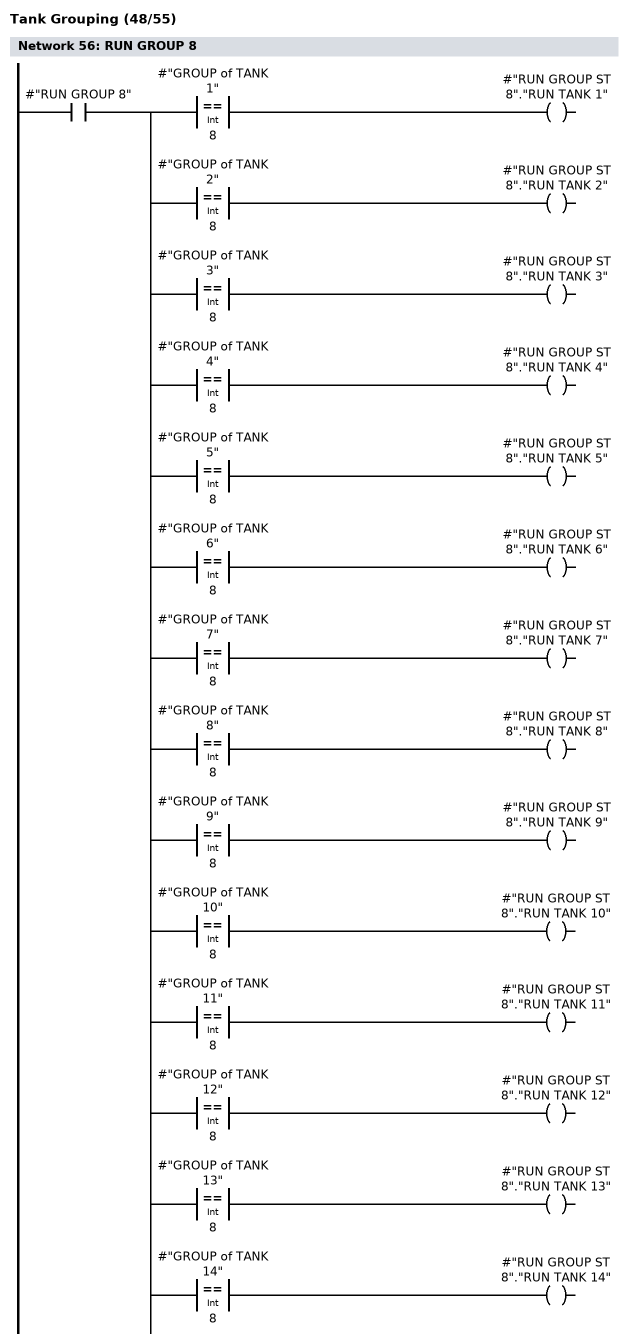
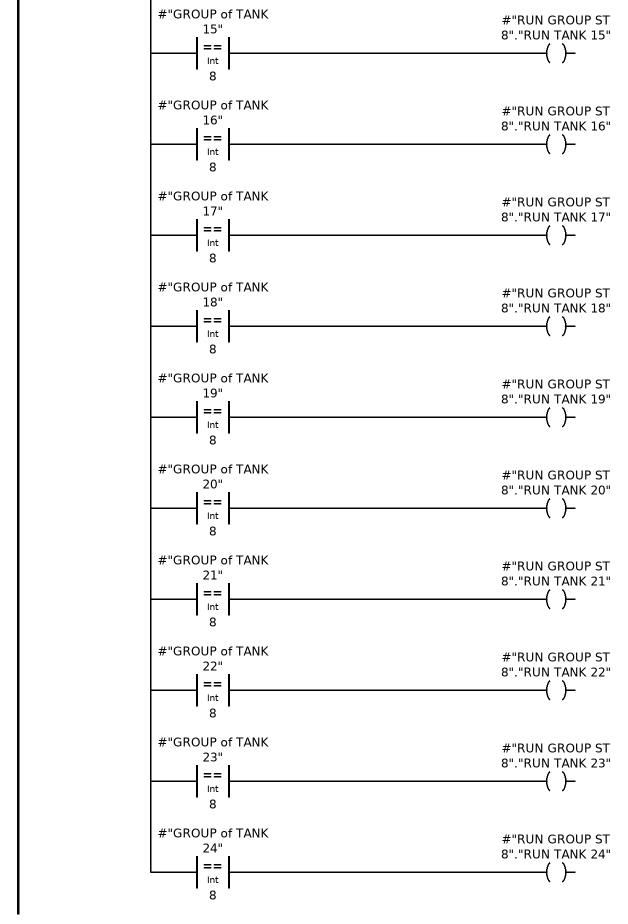
   RUNG wire#powerrail
      Contact( #"RUN GROUP 8" )
      wire#w1
      { S7_Templates := "SrcType := Int" } EQ_Contact(in1 := #"GROUP of TANK 1", in2 := 8)
      Coil( #"RUN GROUP ST 8"."RUN TANK 1" )
   END_RUNG
   RUNG wire#w1
      { S7_Templates := "SrcType := Int" } EQ_Contact(in1 := #"GROUP of TANK 2", in2 := 8)
      Coil( #"RUN GROUP ST 8"."RUN TANK 2" )
   END_RUNG
   RUNG wire#w1
      { S7_Templates := "SrcType := Int" } EQ_Contact(in1 := #"GROUP of TANK 3", in2 := 8)
      Coil( #"RUN GROUP ST 8"."RUN TANK 3" )
   END_RUNG
   RUNG wire#w1
      { S7_Templates := "SrcType := Int" } EQ_Contact(in1 := #"GROUP of TANK 4", in2 := 8)
      Coil( #"RUN GROUP ST 8"."RUN TANK 4" )
   END_RUNG
   RUNG wire#w1
      { S7_Templates := "SrcType := Int" } EQ_Contact(in1 := #"GROUP of TANK 5", in2 := 8)
      Coil( #"RUN GROUP ST 8"."RUN TANK 5" )
   END_RUNG
   RUNG wire#w1
      { S7_Templates := "SrcType := Int" } EQ_Contact(in1 := #"GROUP of TANK 6", in2 := 8)
      Coil( #"RUN GROUP ST 8"."RUN TANK 6" )
   END_RUNG
   RUNG wire#w1
      { S7_Templates := "SrcType := Int" } EQ_Contact(in1 := #"GROUP of TANK 7", in2 := 8)
      Coil( #"RUN GROUP ST 8"."RUN TANK 7" )
   END_RUNG
   RUNG wire#w1
      { S7_Templates := "SrcType := Int" } EQ_Contact(in1 := #"GROUP of TANK 8", in2 := 8)
      Coil( #"RUN GROUP ST 8"."RUN TANK 8" )
   END_RUNG
   RUNG wire#w1
      { S7_Templates := "SrcType := Int" } EQ_Contact(in1 := #"GROUP of TANK 9", in2 := 8)
      Coil( #"RUN GROUP ST 8"."RUN TANK 9" )
   END_RUNG
   RUNG wire#w1
      { S7_Templates := "SrcType := Int" } EQ_Contact(in1 := #"GROUP of TANK 10", in2 := 8)
      Coil( #"RUN GROUP ST 8"."RUN TANK 10" )
   END_RUNG
   RUNG wire#w1
      { S7_Templates := "SrcType := Int" } EQ_Contact(in1 := #"GROUP of TANK 11", in2 := 8)
      Coil( #"RUN GROUP ST 8"."RUN TANK 11" )
   END_RUNG
   RUNG wire#w1
      { S7_Templates := "SrcType := Int" } EQ_Contact(in1 := #"GROUP of TANK 12", in2 := 8)
      Coil( #"RUN GROUP ST 8"."RUN TANK 12" )
   END_RUNG
   RUNG wire#w1
      { S7_Templates := "SrcType := Int" } EQ_Contact(in1 := #"GROUP of TANK 13", in2 := 8)
      Coil( #"RUN GROUP ST 8"."RUN TANK 13" )
   END_RUNG
   RUNG wire#w1
      { S7_Templates := "SrcType := Int" } EQ_Contact(in1 := #"GROUP of TANK 14", in2 := 8)
      Coil( #"RUN GROUP ST 8"."RUN TANK 14" )
   END_RUNG
   RUNG wire#w1
      { S7_Templates := "SrcType := Int" } EQ_Contact(in1 := #"GROUP of TANK 15", in2 := 8)
      Coil( #"RUN GROUP ST 8"."RUN TANK 15" )
   END_RUNG
   RUNG wire#w1
      { S7_Templates := "SrcType := Int" } EQ_Contact(in1 := #"GROUP of TANK 16", in2 := 8)
      Coil( #"RUN GROUP ST 8"."RUN TANK 16" )
   END_RUNG
   RUNG wire#w1
      { S7_Templates := "SrcType := Int" } EQ_Contact(in1 := #"GROUP of TANK 17", in2 := 8)
      Coil( #"RUN GROUP ST 8"."RUN TANK 17" )
   END_RUNG
   RUNG wire#w1
      { S7_Templates := "SrcType := Int" } EQ_Contact(in1 := #"GROUP of TANK 18", in2 := 8)
      Coil( #"RUN GROUP ST 8"."RUN TANK 18" )
   END_RUNG
   RUNG wire#w1
      { S7_Templates := "SrcType := Int" } EQ_Contact(in1 := #"GROUP of TANK 19", in2 := 8)
      Coil( #"RUN GROUP ST 8"."RUN TANK 19" )
   END_RUNG
   RUNG wire#w1
      { S7_Templates := "SrcType := Int" } EQ_Contact(in1 := #"GROUP of TANK 20", in2 := 8)
      Coil( #"RUN GROUP ST 8"."RUN TANK 20" )
   END_RUNG
   RUNG wire#w1
      { S7_Templates := "SrcType := Int" } EQ_Contact(in1 := #"GROUP of TANK 21", in2 := 8)
      Coil( #"RUN GROUP ST 8"."RUN TANK 21" )
   END_RUNG
   RUNG wire#w1
      { S7_Templates := "SrcType := Int" } EQ_Contact(in1 := #"GROUP of TANK 22", in2 := 8)
      Coil( #"RUN GROUP ST 8"."RUN TANK 22" )
   END_RUNG
   RUNG wire#w1
      { S7_Templates := "SrcType := Int" } EQ_Contact(in1 := #"GROUP of TANK 23", in2 := 8)
      Coil( #"RUN GROUP ST 8"."RUN TANK 23" )
   END_RUNG
   RUNG wire#w1
      { S7_Templates := "SrcType := Int" } EQ_Contact(in1 := #"GROUP of TANK 24", in2 := 8)
      Coil( #"RUN GROUP ST 8"."RUN TANK 24" )
   END_RUNG
   // the same network as SCL:
   #"RUN GROUP ST 8"."RUN TANK 1" := #"RUN GROUP 8" AND (#"GROUP of TANK 1" = 8);
   #"RUN GROUP ST 8"."RUN TANK 2" := #"RUN GROUP 8" AND (#"GROUP of TANK 2" = 8);
   #"RUN GROUP ST 8"."RUN TANK 3" := #"RUN GROUP 8" AND (#"GROUP of TANK 3" = 8);
   #"RUN GROUP ST 8"."RUN TANK 4" := #"RUN GROUP 8" AND (#"GROUP of TANK 4" = 8);
   #"RUN GROUP ST 8"."RUN TANK 5" := #"RUN GROUP 8" AND (#"GROUP of TANK 5" = 8);
   #"RUN GROUP ST 8"."RUN TANK 6" := #"RUN GROUP 8" AND (#"GROUP of TANK 6" = 8);
   #"RUN GROUP ST 8"."RUN TANK 7" := #"RUN GROUP 8" AND (#"GROUP of TANK 7" = 8);
   #"RUN GROUP ST 8"."RUN TANK 8" := #"RUN GROUP 8" AND (#"GROUP of TANK 8" = 8);
   #"RUN GROUP ST 8"."RUN TANK 9" := #"RUN GROUP 8" AND (#"GROUP of TANK 9" = 8);
   #"RUN GROUP ST 8"."RUN TANK 10" := #"RUN GROUP 8" AND (#"GROUP of TANK 10" = 8);
   #"RUN GROUP ST 8"."RUN TANK 11" := #"RUN GROUP 8" AND (#"GROUP of TANK 11" = 8);
   #"RUN GROUP ST 8"."RUN TANK 12" := #"RUN GROUP 8" AND (#"GROUP of TANK 12" = 8);
   #"RUN GROUP ST 8"."RUN TANK 13" := #"RUN GROUP 8" AND (#"GROUP of TANK 13" = 8);
   #"RUN GROUP ST 8"."RUN TANK 14" := #"RUN GROUP 8" AND (#"GROUP of TANK 14" = 8);
   #"RUN GROUP ST 8"."RUN TANK 15" := #"RUN GROUP 8" AND (#"GROUP of TANK 15" = 8);
   #"RUN GROUP ST 8"."RUN TANK 16" := #"RUN GROUP 8" AND (#"GROUP of TANK 16" = 8);
   #"RUN GROUP ST 8"."RUN TANK 17" := #"RUN GROUP 8" AND (#"GROUP of TANK 17" = 8);
   #"RUN GROUP ST 8"."RUN TANK 18" := #"RUN GROUP 8" AND (#"GROUP of TANK 18" = 8);
   #"RUN GROUP ST 8"."RUN TANK 19" := #"RUN GROUP 8" AND (#"GROUP of TANK 19" = 8);
   #"RUN GROUP ST 8"."RUN TANK 20" := #"RUN GROUP 8" AND (#"GROUP of TANK 20" = 8);
   #"RUN GROUP ST 8"."RUN TANK 21" := #"RUN GROUP 8" AND (#"GROUP of TANK 21" = 8);
   #"RUN GROUP ST 8"."RUN TANK 22" := #"RUN GROUP 8" AND (#"GROUP of TANK 22" = 8);
   #"RUN GROUP ST 8"."RUN TANK 23" := #"RUN GROUP 8" AND (#"GROUP of TANK 23" = 8);
   #"RUN GROUP ST 8"."RUN TANK 24" := #"RUN GROUP 8" AND (#"GROUP of TANK 24" = 8);
END_REGION

REGION Network 57: RUN GROUP 9
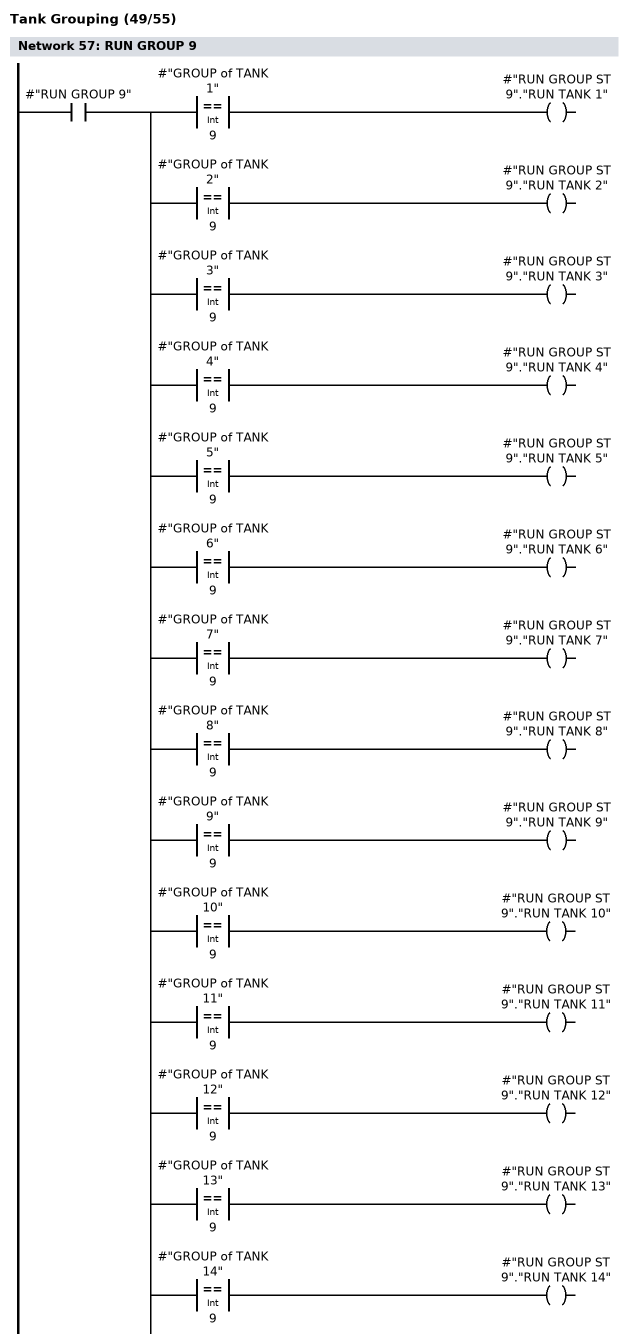
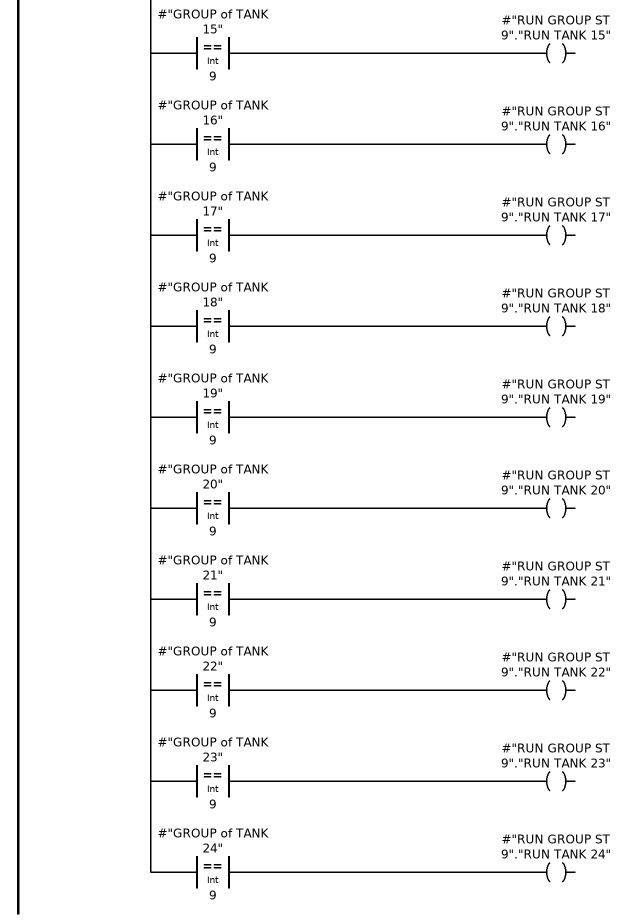
   RUNG wire#powerrail
      Contact( #"RUN GROUP 9" )
      wire#w1
      { S7_Templates := "SrcType := Int" } EQ_Contact(in1 := #"GROUP of TANK 1", in2 := 9)
      Coil( #"RUN GROUP ST 9"."RUN TANK 1" )
   END_RUNG
   RUNG wire#w1
      { S7_Templates := "SrcType := Int" } EQ_Contact(in1 := #"GROUP of TANK 2", in2 := 9)
      Coil( #"RUN GROUP ST 9"."RUN TANK 2" )
   END_RUNG
   RUNG wire#w1
      { S7_Templates := "SrcType := Int" } EQ_Contact(in1 := #"GROUP of TANK 3", in2 := 9)
      Coil( #"RUN GROUP ST 9"."RUN TANK 3" )
   END_RUNG
   RUNG wire#w1
      { S7_Templates := "SrcType := Int" } EQ_Contact(in1 := #"GROUP of TANK 4", in2 := 9)
      Coil( #"RUN GROUP ST 9"."RUN TANK 4" )
   END_RUNG
   RUNG wire#w1
      { S7_Templates := "SrcType := Int" } EQ_Contact(in1 := #"GROUP of TANK 5", in2 := 9)
      Coil( #"RUN GROUP ST 9"."RUN TANK 5" )
   END_RUNG
   RUNG wire#w1
      { S7_Templates := "SrcType := Int" } EQ_Contact(in1 := #"GROUP of TANK 6", in2 := 9)
      Coil( #"RUN GROUP ST 9"."RUN TANK 6" )
   END_RUNG
   RUNG wire#w1
      { S7_Templates := "SrcType := Int" } EQ_Contact(in1 := #"GROUP of TANK 7", in2 := 9)
      Coil( #"RUN GROUP ST 9"."RUN TANK 7" )
   END_RUNG
   RUNG wire#w1
      { S7_Templates := "SrcType := Int" } EQ_Contact(in1 := #"GROUP of TANK 8", in2 := 9)
      Coil( #"RUN GROUP ST 9"."RUN TANK 8" )
   END_RUNG
   RUNG wire#w1
      { S7_Templates := "SrcType := Int" } EQ_Contact(in1 := #"GROUP of TANK 9", in2 := 9)
      Coil( #"RUN GROUP ST 9"."RUN TANK 9" )
   END_RUNG
   RUNG wire#w1
      { S7_Templates := "SrcType := Int" } EQ_Contact(in1 := #"GROUP of TANK 10", in2 := 9)
      Coil( #"RUN GROUP ST 9"."RUN TANK 10" )
   END_RUNG
   RUNG wire#w1
      { S7_Templates := "SrcType := Int" } EQ_Contact(in1 := #"GROUP of TANK 11", in2 := 9)
      Coil( #"RUN GROUP ST 9"."RUN TANK 11" )
   END_RUNG
   RUNG wire#w1
      { S7_Templates := "SrcType := Int" } EQ_Contact(in1 := #"GROUP of TANK 12", in2 := 9)
      Coil( #"RUN GROUP ST 9"."RUN TANK 12" )
   END_RUNG
   RUNG wire#w1
      { S7_Templates := "SrcType := Int" } EQ_Contact(in1 := #"GROUP of TANK 13", in2 := 9)
      Coil( #"RUN GROUP ST 9"."RUN TANK 13" )
   END_RUNG
   RUNG wire#w1
      { S7_Templates := "SrcType := Int" } EQ_Contact(in1 := #"GROUP of TANK 14", in2 := 9)
      Coil( #"RUN GROUP ST 9"."RUN TANK 14" )
   END_RUNG
   RUNG wire#w1
      { S7_Templates := "SrcType := Int" } EQ_Contact(in1 := #"GROUP of TANK 15", in2 := 9)
      Coil( #"RUN GROUP ST 9"."RUN TANK 15" )
   END_RUNG
   RUNG wire#w1
      { S7_Templates := "SrcType := Int" } EQ_Contact(in1 := #"GROUP of TANK 16", in2 := 9)
      Coil( #"RUN GROUP ST 9"."RUN TANK 16" )
   END_RUNG
   RUNG wire#w1
      { S7_Templates := "SrcType := Int" } EQ_Contact(in1 := #"GROUP of TANK 17", in2 := 9)
      Coil( #"RUN GROUP ST 9"."RUN TANK 17" )
   END_RUNG
   RUNG wire#w1
      { S7_Templates := "SrcType := Int" } EQ_Contact(in1 := #"GROUP of TANK 18", in2 := 9)
      Coil( #"RUN GROUP ST 9"."RUN TANK 18" )
   END_RUNG
   RUNG wire#w1
      { S7_Templates := "SrcType := Int" } EQ_Contact(in1 := #"GROUP of TANK 19", in2 := 9)
      Coil( #"RUN GROUP ST 9"."RUN TANK 19" )
   END_RUNG
   RUNG wire#w1
      { S7_Templates := "SrcType := Int" } EQ_Contact(in1 := #"GROUP of TANK 20", in2 := 9)
      Coil( #"RUN GROUP ST 9"."RUN TANK 20" )
   END_RUNG
   RUNG wire#w1
      { S7_Templates := "SrcType := Int" } EQ_Contact(in1 := #"GROUP of TANK 21", in2 := 9)
      Coil( #"RUN GROUP ST 9"."RUN TANK 21" )
   END_RUNG
   RUNG wire#w1
      { S7_Templates := "SrcType := Int" } EQ_Contact(in1 := #"GROUP of TANK 22", in2 := 9)
      Coil( #"RUN GROUP ST 9"."RUN TANK 22" )
   END_RUNG
   RUNG wire#w1
      { S7_Templates := "SrcType := Int" } EQ_Contact(in1 := #"GROUP of TANK 23", in2 := 9)
      Coil( #"RUN GROUP ST 9"."RUN TANK 23" )
   END_RUNG
   RUNG wire#w1
      { S7_Templates := "SrcType := Int" } EQ_Contact(in1 := #"GROUP of TANK 24", in2 := 9)
      Coil( #"RUN GROUP ST 9"."RUN TANK 24" )
   END_RUNG
   // the same network as SCL:
   #"RUN GROUP ST 9"."RUN TANK 1" := #"RUN GROUP 9" AND (#"GROUP of TANK 1" = 9);
   #"RUN GROUP ST 9"."RUN TANK 2" := #"RUN GROUP 9" AND (#"GROUP of TANK 2" = 9);
   #"RUN GROUP ST 9"."RUN TANK 3" := #"RUN GROUP 9" AND (#"GROUP of TANK 3" = 9);
   #"RUN GROUP ST 9"."RUN TANK 4" := #"RUN GROUP 9" AND (#"GROUP of TANK 4" = 9);
   #"RUN GROUP ST 9"."RUN TANK 5" := #"RUN GROUP 9" AND (#"GROUP of TANK 5" = 9);
   #"RUN GROUP ST 9"."RUN TANK 6" := #"RUN GROUP 9" AND (#"GROUP of TANK 6" = 9);
   #"RUN GROUP ST 9"."RUN TANK 7" := #"RUN GROUP 9" AND (#"GROUP of TANK 7" = 9);
   #"RUN GROUP ST 9"."RUN TANK 8" := #"RUN GROUP 9" AND (#"GROUP of TANK 8" = 9);
   #"RUN GROUP ST 9"."RUN TANK 9" := #"RUN GROUP 9" AND (#"GROUP of TANK 9" = 9);
   #"RUN GROUP ST 9"."RUN TANK 10" := #"RUN GROUP 9" AND (#"GROUP of TANK 10" = 9);
   #"RUN GROUP ST 9"."RUN TANK 11" := #"RUN GROUP 9" AND (#"GROUP of TANK 11" = 9);
   #"RUN GROUP ST 9"."RUN TANK 12" := #"RUN GROUP 9" AND (#"GROUP of TANK 12" = 9);
   #"RUN GROUP ST 9"."RUN TANK 13" := #"RUN GROUP 9" AND (#"GROUP of TANK 13" = 9);
   #"RUN GROUP ST 9"."RUN TANK 14" := #"RUN GROUP 9" AND (#"GROUP of TANK 14" = 9);
   #"RUN GROUP ST 9"."RUN TANK 15" := #"RUN GROUP 9" AND (#"GROUP of TANK 15" = 9);
   #"RUN GROUP ST 9"."RUN TANK 16" := #"RUN GROUP 9" AND (#"GROUP of TANK 16" = 9);
   #"RUN GROUP ST 9"."RUN TANK 17" := #"RUN GROUP 9" AND (#"GROUP of TANK 17" = 9);
   #"RUN GROUP ST 9"."RUN TANK 18" := #"RUN GROUP 9" AND (#"GROUP of TANK 18" = 9);
   #"RUN GROUP ST 9"."RUN TANK 19" := #"RUN GROUP 9" AND (#"GROUP of TANK 19" = 9);
   #"RUN GROUP ST 9"."RUN TANK 20" := #"RUN GROUP 9" AND (#"GROUP of TANK 20" = 9);
   #"RUN GROUP ST 9"."RUN TANK 21" := #"RUN GROUP 9" AND (#"GROUP of TANK 21" = 9);
   #"RUN GROUP ST 9"."RUN TANK 22" := #"RUN GROUP 9" AND (#"GROUP of TANK 22" = 9);
   #"RUN GROUP ST 9"."RUN TANK 23" := #"RUN GROUP 9" AND (#"GROUP of TANK 23" = 9);
   #"RUN GROUP ST 9"."RUN TANK 24" := #"RUN GROUP 9" AND (#"GROUP of TANK 24" = 9);
END_REGION

REGION Network 58: RUN GROUP 10
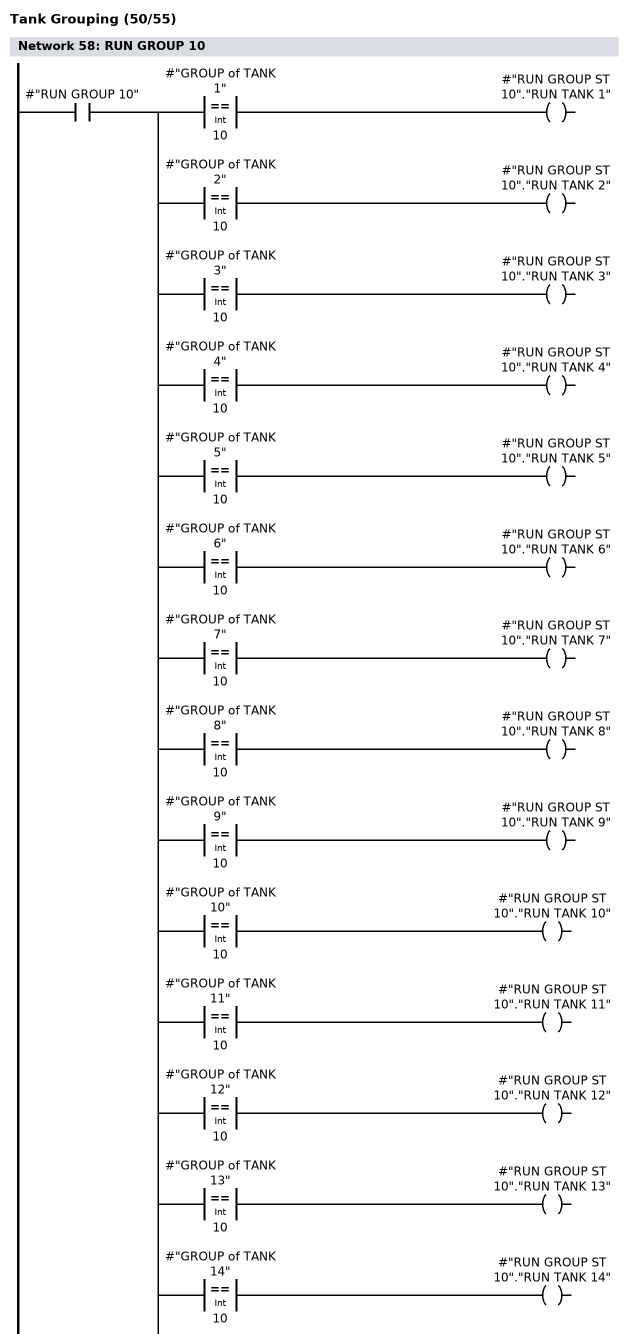
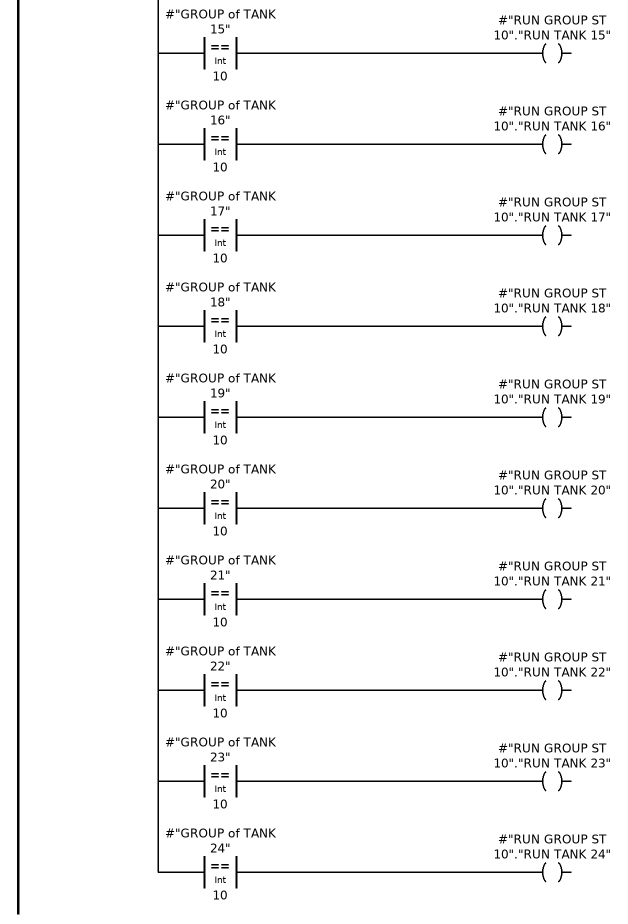
   RUNG wire#powerrail
      Contact( #"RUN GROUP 10" )
      wire#w1
      { S7_Templates := "SrcType := Int" } EQ_Contact(in1 := #"GROUP of TANK 1", in2 := 10)
      Coil( #"RUN GROUP ST 10"."RUN TANK 1" )
   END_RUNG
   RUNG wire#w1
      { S7_Templates := "SrcType := Int" } EQ_Contact(in1 := #"GROUP of TANK 2", in2 := 10)
      Coil( #"RUN GROUP ST 10"."RUN TANK 2" )
   END_RUNG
   RUNG wire#w1
      { S7_Templates := "SrcType := Int" } EQ_Contact(in1 := #"GROUP of TANK 3", in2 := 10)
      Coil( #"RUN GROUP ST 10"."RUN TANK 3" )
   END_RUNG
   RUNG wire#w1
      { S7_Templates := "SrcType := Int" } EQ_Contact(in1 := #"GROUP of TANK 4", in2 := 10)
      Coil( #"RUN GROUP ST 10"."RUN TANK 4" )
   END_RUNG
   RUNG wire#w1
      { S7_Templates := "SrcType := Int" } EQ_Contact(in1 := #"GROUP of TANK 5", in2 := 10)
      Coil( #"RUN GROUP ST 10"."RUN TANK 5" )
   END_RUNG
   RUNG wire#w1
      { S7_Templates := "SrcType := Int" } EQ_Contact(in1 := #"GROUP of TANK 6", in2 := 10)
      Coil( #"RUN GROUP ST 10"."RUN TANK 6" )
   END_RUNG
   RUNG wire#w1
      { S7_Templates := "SrcType := Int" } EQ_Contact(in1 := #"GROUP of TANK 7", in2 := 10)
      Coil( #"RUN GROUP ST 10"."RUN TANK 7" )
   END_RUNG
   RUNG wire#w1
      { S7_Templates := "SrcType := Int" } EQ_Contact(in1 := #"GROUP of TANK 8", in2 := 10)
      Coil( #"RUN GROUP ST 10"."RUN TANK 8" )
   END_RUNG
   RUNG wire#w1
      { S7_Templates := "SrcType := Int" } EQ_Contact(in1 := #"GROUP of TANK 9", in2 := 10)
      Coil( #"RUN GROUP ST 10"."RUN TANK 9" )
   END_RUNG
   RUNG wire#w1
      { S7_Templates := "SrcType := Int" } EQ_Contact(in1 := #"GROUP of TANK 10", in2 := 10)
      Coil( #"RUN GROUP ST 10"."RUN TANK 10" )
   END_RUNG
   RUNG wire#w1
      { S7_Templates := "SrcType := Int" } EQ_Contact(in1 := #"GROUP of TANK 11", in2 := 10)
      Coil( #"RUN GROUP ST 10"."RUN TANK 11" )
   END_RUNG
   RUNG wire#w1
      { S7_Templates := "SrcType := Int" } EQ_Contact(in1 := #"GROUP of TANK 12", in2 := 10)
      Coil( #"RUN GROUP ST 10"."RUN TANK 12" )
   END_RUNG
   RUNG wire#w1
      { S7_Templates := "SrcType := Int" } EQ_Contact(in1 := #"GROUP of TANK 13", in2 := 10)
      Coil( #"RUN GROUP ST 10"."RUN TANK 13" )
   END_RUNG
   RUNG wire#w1
      { S7_Templates := "SrcType := Int" } EQ_Contact(in1 := #"GROUP of TANK 14", in2 := 10)
      Coil( #"RUN GROUP ST 10"."RUN TANK 14" )
   END_RUNG
   RUNG wire#w1
      { S7_Templates := "SrcType := Int" } EQ_Contact(in1 := #"GROUP of TANK 15", in2 := 10)
      Coil( #"RUN GROUP ST 10"."RUN TANK 15" )
   END_RUNG
   RUNG wire#w1
      { S7_Templates := "SrcType := Int" } EQ_Contact(in1 := #"GROUP of TANK 16", in2 := 10)
      Coil( #"RUN GROUP ST 10"."RUN TANK 16" )
   END_RUNG
   RUNG wire#w1
      { S7_Templates := "SrcType := Int" } EQ_Contact(in1 := #"GROUP of TANK 17", in2 := 10)
      Coil( #"RUN GROUP ST 10"."RUN TANK 17" )
   END_RUNG
   RUNG wire#w1
      { S7_Templates := "SrcType := Int" } EQ_Contact(in1 := #"GROUP of TANK 18", in2 := 10)
      Coil( #"RUN GROUP ST 10"."RUN TANK 18" )
   END_RUNG
   RUNG wire#w1
      { S7_Templates := "SrcType := Int" } EQ_Contact(in1 := #"GROUP of TANK 19", in2 := 10)
      Coil( #"RUN GROUP ST 10"."RUN TANK 19" )
   END_RUNG
   RUNG wire#w1
      { S7_Templates := "SrcType := Int" } EQ_Contact(in1 := #"GROUP of TANK 20", in2 := 10)
      Coil( #"RUN GROUP ST 10"."RUN TANK 20" )
   END_RUNG
   RUNG wire#w1
      { S7_Templates := "SrcType := Int" } EQ_Contact(in1 := #"GROUP of TANK 21", in2 := 10)
      Coil( #"RUN GROUP ST 10"."RUN TANK 21" )
   END_RUNG
   RUNG wire#w1
      { S7_Templates := "SrcType := Int" } EQ_Contact(in1 := #"GROUP of TANK 22", in2 := 10)
      Coil( #"RUN GROUP ST 10"."RUN TANK 22" )
   END_RUNG
   RUNG wire#w1
      { S7_Templates := "SrcType := Int" } EQ_Contact(in1 := #"GROUP of TANK 23", in2 := 10)
      Coil( #"RUN GROUP ST 10"."RUN TANK 23" )
   END_RUNG
   RUNG wire#w1
      { S7_Templates := "SrcType := Int" } EQ_Contact(in1 := #"GROUP of TANK 24", in2 := 10)
      Coil( #"RUN GROUP ST 10"."RUN TANK 24" )
   END_RUNG
   // the same network as SCL:
   #"RUN GROUP ST 10"."RUN TANK 1" := #"RUN GROUP 10" AND (#"GROUP of TANK 1" = 10);
   #"RUN GROUP ST 10"."RUN TANK 2" := #"RUN GROUP 10" AND (#"GROUP of TANK 2" = 10);
   #"RUN GROUP ST 10"."RUN TANK 3" := #"RUN GROUP 10" AND (#"GROUP of TANK 3" = 10);
   #"RUN GROUP ST 10"."RUN TANK 4" := #"RUN GROUP 10" AND (#"GROUP of TANK 4" = 10);
   #"RUN GROUP ST 10"."RUN TANK 5" := #"RUN GROUP 10" AND (#"GROUP of TANK 5" = 10);
   #"RUN GROUP ST 10"."RUN TANK 6" := #"RUN GROUP 10" AND (#"GROUP of TANK 6" = 10);
   #"RUN GROUP ST 10"."RUN TANK 7" := #"RUN GROUP 10" AND (#"GROUP of TANK 7" = 10);
   #"RUN GROUP ST 10"."RUN TANK 8" := #"RUN GROUP 10" AND (#"GROUP of TANK 8" = 10);
   #"RUN GROUP ST 10"."RUN TANK 9" := #"RUN GROUP 10" AND (#"GROUP of TANK 9" = 10);
   #"RUN GROUP ST 10"."RUN TANK 10" := #"RUN GROUP 10" AND (#"GROUP of TANK 10" = 10);
   #"RUN GROUP ST 10"."RUN TANK 11" := #"RUN GROUP 10" AND (#"GROUP of TANK 11" = 10);
   #"RUN GROUP ST 10"."RUN TANK 12" := #"RUN GROUP 10" AND (#"GROUP of TANK 12" = 10);
   #"RUN GROUP ST 10"."RUN TANK 13" := #"RUN GROUP 10" AND (#"GROUP of TANK 13" = 10);
   #"RUN GROUP ST 10"."RUN TANK 14" := #"RUN GROUP 10" AND (#"GROUP of TANK 14" = 10);
   #"RUN GROUP ST 10"."RUN TANK 15" := #"RUN GROUP 10" AND (#"GROUP of TANK 15" = 10);
   #"RUN GROUP ST 10"."RUN TANK 16" := #"RUN GROUP 10" AND (#"GROUP of TANK 16" = 10);
   #"RUN GROUP ST 10"."RUN TANK 17" := #"RUN GROUP 10" AND (#"GROUP of TANK 17" = 10);
   #"RUN GROUP ST 10"."RUN TANK 18" := #"RUN GROUP 10" AND (#"GROUP of TANK 18" = 10);
   #"RUN GROUP ST 10"."RUN TANK 19" := #"RUN GROUP 10" AND (#"GROUP of TANK 19" = 10);
   #"RUN GROUP ST 10"."RUN TANK 20" := #"RUN GROUP 10" AND (#"GROUP of TANK 20" = 10);
   #"RUN GROUP ST 10"."RUN TANK 21" := #"RUN GROUP 10" AND (#"GROUP of TANK 21" = 10);
   #"RUN GROUP ST 10"."RUN TANK 22" := #"RUN GROUP 10" AND (#"GROUP of TANK 22" = 10);
   #"RUN GROUP ST 10"."RUN TANK 23" := #"RUN GROUP 10" AND (#"GROUP of TANK 23" = 10);
   #"RUN GROUP ST 10"."RUN TANK 24" := #"RUN GROUP 10" AND (#"GROUP of TANK 24" = 10);
END_REGION

REGION Network 59: RUN GROUP 11
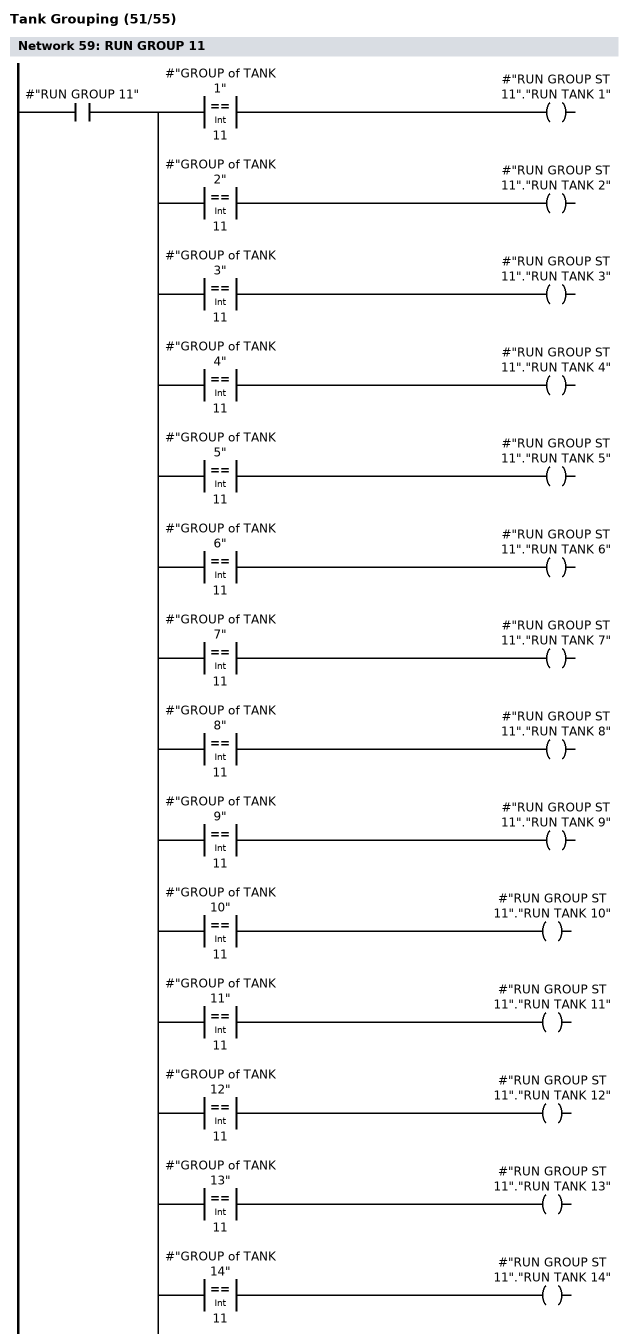
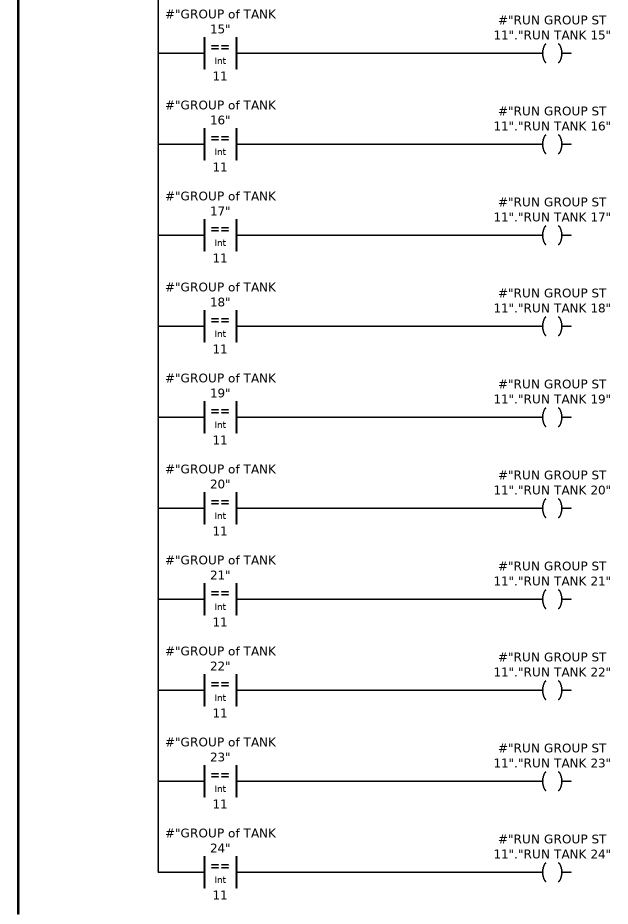
   RUNG wire#powerrail
      Contact( #"RUN GROUP 11" )
      wire#w1
      { S7_Templates := "SrcType := Int" } EQ_Contact(in1 := #"GROUP of TANK 1", in2 := 11)
      Coil( #"RUN GROUP ST 11"."RUN TANK 1" )
   END_RUNG
   RUNG wire#w1
      { S7_Templates := "SrcType := Int" } EQ_Contact(in1 := #"GROUP of TANK 2", in2 := 11)
      Coil( #"RUN GROUP ST 11"."RUN TANK 2" )
   END_RUNG
   RUNG wire#w1
      { S7_Templates := "SrcType := Int" } EQ_Contact(in1 := #"GROUP of TANK 3", in2 := 11)
      Coil( #"RUN GROUP ST 11"."RUN TANK 3" )
   END_RUNG
   RUNG wire#w1
      { S7_Templates := "SrcType := Int" } EQ_Contact(in1 := #"GROUP of TANK 4", in2 := 11)
      Coil( #"RUN GROUP ST 11"."RUN TANK 4" )
   END_RUNG
   RUNG wire#w1
      { S7_Templates := "SrcType := Int" } EQ_Contact(in1 := #"GROUP of TANK 5", in2 := 11)
      Coil( #"RUN GROUP ST 11"."RUN TANK 5" )
   END_RUNG
   RUNG wire#w1
      { S7_Templates := "SrcType := Int" } EQ_Contact(in1 := #"GROUP of TANK 6", in2 := 11)
      Coil( #"RUN GROUP ST 11"."RUN TANK 6" )
   END_RUNG
   RUNG wire#w1
      { S7_Templates := "SrcType := Int" } EQ_Contact(in1 := #"GROUP of TANK 7", in2 := 11)
      Coil( #"RUN GROUP ST 11"."RUN TANK 7" )
   END_RUNG
   RUNG wire#w1
      { S7_Templates := "SrcType := Int" } EQ_Contact(in1 := #"GROUP of TANK 8", in2 := 11)
      Coil( #"RUN GROUP ST 11"."RUN TANK 8" )
   END_RUNG
   RUNG wire#w1
      { S7_Templates := "SrcType := Int" } EQ_Contact(in1 := #"GROUP of TANK 9", in2 := 11)
      Coil( #"RUN GROUP ST 11"."RUN TANK 9" )
   END_RUNG
   RUNG wire#w1
      { S7_Templates := "SrcType := Int" } EQ_Contact(in1 := #"GROUP of TANK 10", in2 := 11)
      Coil( #"RUN GROUP ST 11"."RUN TANK 10" )
   END_RUNG
   RUNG wire#w1
      { S7_Templates := "SrcType := Int" } EQ_Contact(in1 := #"GROUP of TANK 11", in2 := 11)
      Coil( #"RUN GROUP ST 11"."RUN TANK 11" )
   END_RUNG
   RUNG wire#w1
      { S7_Templates := "SrcType := Int" } EQ_Contact(in1 := #"GROUP of TANK 12", in2 := 11)
      Coil( #"RUN GROUP ST 11"."RUN TANK 12" )
   END_RUNG
   RUNG wire#w1
      { S7_Templates := "SrcType := Int" } EQ_Contact(in1 := #"GROUP of TANK 13", in2 := 11)
      Coil( #"RUN GROUP ST 11"."RUN TANK 13" )
   END_RUNG
   RUNG wire#w1
      { S7_Templates := "SrcType := Int" } EQ_Contact(in1 := #"GROUP of TANK 14", in2 := 11)
      Coil( #"RUN GROUP ST 11"."RUN TANK 14" )
   END_RUNG
   RUNG wire#w1
      { S7_Templates := "SrcType := Int" } EQ_Contact(in1 := #"GROUP of TANK 15", in2 := 11)
      Coil( #"RUN GROUP ST 11"."RUN TANK 15" )
   END_RUNG
   RUNG wire#w1
      { S7_Templates := "SrcType := Int" } EQ_Contact(in1 := #"GROUP of TANK 16", in2 := 11)
      Coil( #"RUN GROUP ST 11"."RUN TANK 16" )
   END_RUNG
   RUNG wire#w1
      { S7_Templates := "SrcType := Int" } EQ_Contact(in1 := #"GROUP of TANK 17", in2 := 11)
      Coil( #"RUN GROUP ST 11"."RUN TANK 17" )
   END_RUNG
   RUNG wire#w1
      { S7_Templates := "SrcType := Int" } EQ_Contact(in1 := #"GROUP of TANK 18", in2 := 11)
      Coil( #"RUN GROUP ST 11"."RUN TANK 18" )
   END_RUNG
   RUNG wire#w1
      { S7_Templates := "SrcType := Int" } EQ_Contact(in1 := #"GROUP of TANK 19", in2 := 11)
      Coil( #"RUN GROUP ST 11"."RUN TANK 19" )
   END_RUNG
   RUNG wire#w1
      { S7_Templates := "SrcType := Int" } EQ_Contact(in1 := #"GROUP of TANK 20", in2 := 11)
      Coil( #"RUN GROUP ST 11"."RUN TANK 20" )
   END_RUNG
   RUNG wire#w1
      { S7_Templates := "SrcType := Int" } EQ_Contact(in1 := #"GROUP of TANK 21", in2 := 11)
      Coil( #"RUN GROUP ST 11"."RUN TANK 21" )
   END_RUNG
   RUNG wire#w1
      { S7_Templates := "SrcType := Int" } EQ_Contact(in1 := #"GROUP of TANK 22", in2 := 11)
      Coil( #"RUN GROUP ST 11"."RUN TANK 22" )
   END_RUNG
   RUNG wire#w1
      { S7_Templates := "SrcType := Int" } EQ_Contact(in1 := #"GROUP of TANK 23", in2 := 11)
      Coil( #"RUN GROUP ST 11"."RUN TANK 23" )
   END_RUNG
   RUNG wire#w1
      { S7_Templates := "SrcType := Int" } EQ_Contact(in1 := #"GROUP of TANK 24", in2 := 11)
      Coil( #"RUN GROUP ST 11"."RUN TANK 24" )
   END_RUNG
   // the same network as SCL:
   #"RUN GROUP ST 11"."RUN TANK 1" := #"RUN GROUP 11" AND (#"GROUP of TANK 1" = 11);
   #"RUN GROUP ST 11"."RUN TANK 2" := #"RUN GROUP 11" AND (#"GROUP of TANK 2" = 11);
   #"RUN GROUP ST 11"."RUN TANK 3" := #"RUN GROUP 11" AND (#"GROUP of TANK 3" = 11);
   #"RUN GROUP ST 11"."RUN TANK 4" := #"RUN GROUP 11" AND (#"GROUP of TANK 4" = 11);
   #"RUN GROUP ST 11"."RUN TANK 5" := #"RUN GROUP 11" AND (#"GROUP of TANK 5" = 11);
   #"RUN GROUP ST 11"."RUN TANK 6" := #"RUN GROUP 11" AND (#"GROUP of TANK 6" = 11);
   #"RUN GROUP ST 11"."RUN TANK 7" := #"RUN GROUP 11" AND (#"GROUP of TANK 7" = 11);
   #"RUN GROUP ST 11"."RUN TANK 8" := #"RUN GROUP 11" AND (#"GROUP of TANK 8" = 11);
   #"RUN GROUP ST 11"."RUN TANK 9" := #"RUN GROUP 11" AND (#"GROUP of TANK 9" = 11);
   #"RUN GROUP ST 11"."RUN TANK 10" := #"RUN GROUP 11" AND (#"GROUP of TANK 10" = 11);
   #"RUN GROUP ST 11"."RUN TANK 11" := #"RUN GROUP 11" AND (#"GROUP of TANK 11" = 11);
   #"RUN GROUP ST 11"."RUN TANK 12" := #"RUN GROUP 11" AND (#"GROUP of TANK 12" = 11);
   #"RUN GROUP ST 11"."RUN TANK 13" := #"RUN GROUP 11" AND (#"GROUP of TANK 13" = 11);
   #"RUN GROUP ST 11"."RUN TANK 14" := #"RUN GROUP 11" AND (#"GROUP of TANK 14" = 11);
   #"RUN GROUP ST 11"."RUN TANK 15" := #"RUN GROUP 11" AND (#"GROUP of TANK 15" = 11);
   #"RUN GROUP ST 11"."RUN TANK 16" := #"RUN GROUP 11" AND (#"GROUP of TANK 16" = 11);
   #"RUN GROUP ST 11"."RUN TANK 17" := #"RUN GROUP 11" AND (#"GROUP of TANK 17" = 11);
   #"RUN GROUP ST 11"."RUN TANK 18" := #"RUN GROUP 11" AND (#"GROUP of TANK 18" = 11);
   #"RUN GROUP ST 11"."RUN TANK 19" := #"RUN GROUP 11" AND (#"GROUP of TANK 19" = 11);
   #"RUN GROUP ST 11"."RUN TANK 20" := #"RUN GROUP 11" AND (#"GROUP of TANK 20" = 11);
   #"RUN GROUP ST 11"."RUN TANK 21" := #"RUN GROUP 11" AND (#"GROUP of TANK 21" = 11);
   #"RUN GROUP ST 11"."RUN TANK 22" := #"RUN GROUP 11" AND (#"GROUP of TANK 22" = 11);
   #"RUN GROUP ST 11"."RUN TANK 23" := #"RUN GROUP 11" AND (#"GROUP of TANK 23" = 11);
   #"RUN GROUP ST 11"."RUN TANK 24" := #"RUN GROUP 11" AND (#"GROUP of TANK 24" = 11);
END_REGION

REGION Network 60: RUN GROUP 12